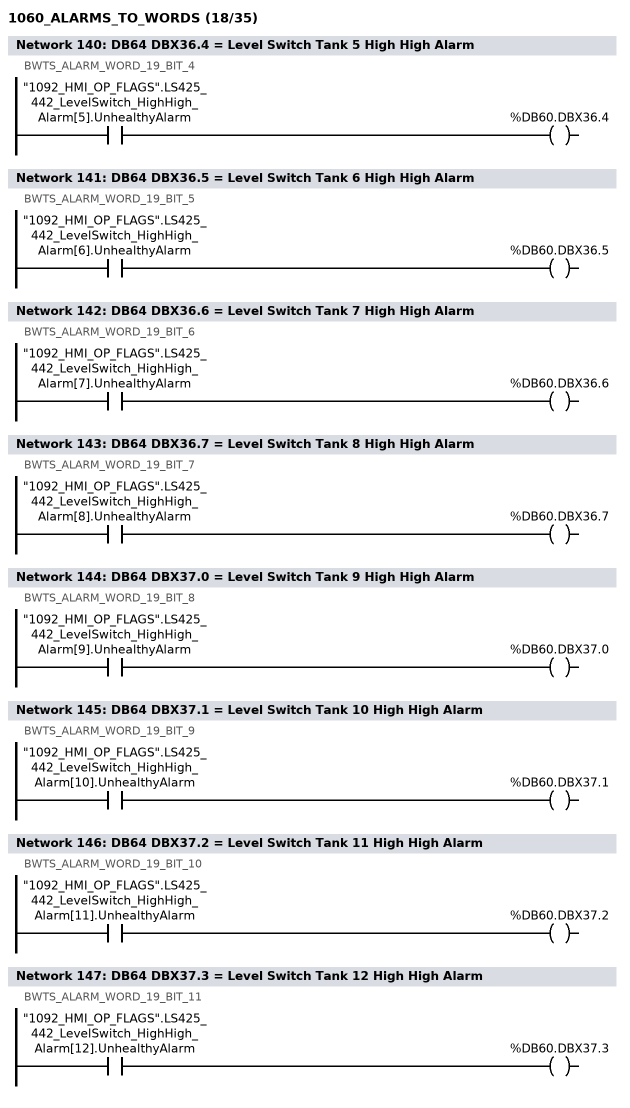
   RUNG wire#powerrail
      Contact( "1092_HMI_OP_FLAGS".LS425_442_LevelSwitch_HighHigh_Alarm[5].UnhealthyAlarm )
      Coil( %DB60.DBX36.4 )
   END_RUNG
   // the same network as SCL:
   %DB60.DBX36.4 := "1092_HMI_OP_FLAGS".LS425_442_LevelSwitch_HighHigh_Alarm[5].UnhealthyAlarm;
END_REGION

REGION Network 141: DB64 DBX36.5 = Level Switch Tank 6 High High Alarm
   // BWTS_ALARM_WORD_19_BIT_5
   RUNG wire#powerrail
      Contact( "1092_HMI_OP_FLAGS".LS425_442_LevelSwitch_HighHigh_Alarm[6].UnhealthyAlarm )
      Coil( %DB60.DBX36.5 )
   END_RUNG
   // the same network as SCL:
   %DB60.DBX36.5 := "1092_HMI_OP_FLAGS".LS425_442_LevelSwitch_HighHigh_Alarm[6].UnhealthyAlarm;
END_REGION

REGION Network 142: DB64 DBX36.6 = Level Switch Tank 7 High High Alarm
   // BWTS_ALARM_WORD_19_BIT_6
   RUNG wire#powerrail
      Contact( "1092_HMI_OP_FLAGS".LS425_442_LevelSwitch_HighHigh_Alarm[7].UnhealthyAlarm )
      Coil( %DB60.DBX36.6 )
   END_RUNG
   // the same network as SCL:
   %DB60.DBX36.6 := "1092_HMI_OP_FLAGS".LS425_442_LevelSwitch_HighHigh_Alarm[7].UnhealthyAlarm;
END_REGION

REGION Network 143: DB64 DBX36.7 = Level Switch Tank 8 High High Alarm
   // BWTS_ALARM_WORD_19_BIT_7
   RUNG wire#powerrail
      Contact( "1092_HMI_OP_FLAGS".LS425_442_LevelSwitch_HighHigh_Alarm[8].UnhealthyAlarm )
      Coil( %DB60.DBX36.7 )
   END_RUNG
   // the same network as SCL:
   %DB60.DBX36.7 := "1092_HMI_OP_FLAGS".LS425_442_LevelSwitch_HighHigh_Alarm[8].UnhealthyAlarm;
END_REGION

REGION Network 144: DB64 DBX37.0 = Level Switch Tank 9 High High Alarm
   // BWTS_ALARM_WORD_19_BIT_8
   RUNG wire#powerrail
      Contact( "1092_HMI_OP_FLAGS".LS425_442_LevelSwitch_HighHigh_Alarm[9].UnhealthyAlarm )
      Coil( %DB60.DBX37.0 )
   END_RUNG
   // the same network as SCL:
   %DB60.DBX37.0 := "1092_HMI_OP_FLAGS".LS425_442_LevelSwitch_HighHigh_Alarm[9].UnhealthyAlarm;
END_REGION

REGION Network 145: DB64 DBX37.1 = Level Switch Tank 10 High High Alarm
   // BWTS_ALARM_WORD_19_BIT_9
   RUNG wire#powerrail
      Contact( "1092_HMI_OP_FLAGS".LS425_442_LevelSwitch_HighHigh_Alarm[10].UnhealthyAlarm )
      Coil( %DB60.DBX37.1 )
   END_RUNG
   // the same network as SCL:
   %DB60.DBX37.1 := "1092_HMI_OP_FLAGS".LS425_442_LevelSwitch_HighHigh_Alarm[10].UnhealthyAlarm;
END_REGION

REGION Network 146: DB64 DBX37.2 = Level Switch Tank 11 High High Alarm
   // BWTS_ALARM_WORD_19_BIT_10
   RUNG wire#powerrail
      Contact( "1092_HMI_OP_FLAGS".LS425_442_LevelSwitch_HighHigh_Alarm[11].UnhealthyAlarm )
      Coil( %DB60.DBX37.2 )
   END_RUNG
   // the same network as SCL:
   %DB60.DBX37.2 := "1092_HMI_OP_FLAGS".LS425_442_LevelSwitch_HighHigh_Alarm[11].UnhealthyAlarm;
END_REGION

REGION Network 147: DB64 DBX37.3 = Level Switch Tank 12 High High Alarm
   // BWTS_ALARM_WORD_19_BIT_11
   RUNG wire#powerrail
      Contact( "1092_HMI_OP_FLAGS".LS425_442_LevelSwitch_HighHigh_Alarm[12].UnhealthyAlarm )
      Coil( %DB60.DBX37.3 )
   END_RUNG
   // the same network as SCL:
   %DB60.DBX37.3 := "1092_HMI_OP_FLAGS".LS425_442_LevelSwitch_HighHigh_Alarm[12].UnhealthyAlarm;
END_REGION

REGION Network 148: DB64 DBX37.4 = Level Switch Tank 13 High High Alarm
   // BWTS_ALARM_WORD_19_BIT_12
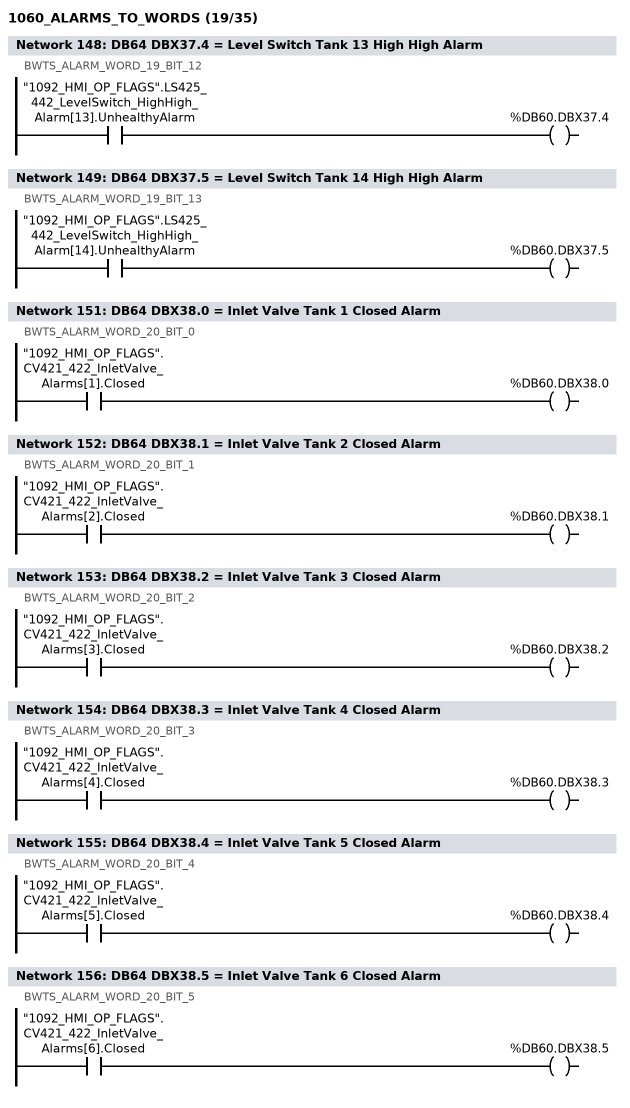
   RUNG wire#powerrail
      Contact( "1092_HMI_OP_FLAGS".LS425_442_LevelSwitch_HighHigh_Alarm[13].UnhealthyAlarm )
      Coil( %DB60.DBX37.4 )
   END_RUNG
   // the same network as SCL:
   %DB60.DBX37.4 := "1092_HMI_OP_FLAGS".LS425_442_LevelSwitch_HighHigh_Alarm[13].UnhealthyAlarm;
END_REGION

REGION Network 149: DB64 DBX37.5 = Level Switch Tank 14 High High Alarm
   // BWTS_ALARM_WORD_19_BIT_13
   RUNG wire#powerrail
      Contact( "1092_HMI_OP_FLAGS".LS425_442_LevelSwitch_HighHigh_Alarm[14].UnhealthyAlarm )
      Coil( %DB60.DBX37.5 )
   END_RUNG
   // the same network as SCL:
   %DB60.DBX37.5 := "1092_HMI_OP_FLAGS".LS425_442_LevelSwitch_HighHigh_Alarm[14].UnhealthyAlarm;
END_REGION

REGION Network 151: DB64 DBX38.0 = Inlet Valve Tank 1 Closed Alarm
   // BWTS_ALARM_WORD_20_BIT_0
   RUNG wire#powerrail
      Contact( "1092_HMI_OP_FLAGS".CV421_422_InletValve_Alarms[1].Closed )
      Coil( %DB60.DBX38.0 )
   END_RUNG
   // the same network as SCL:
   %DB60.DBX38.0 := "1092_HMI_OP_FLAGS".CV421_422_InletValve_Alarms[1].Closed;
END_REGION

REGION Network 152: DB64 DBX38.1 = Inlet Valve Tank 2 Closed Alarm
   // BWTS_ALARM_WORD_20_BIT_1
   RUNG wire#powerrail
      Contact( "1092_HMI_OP_FLAGS".CV421_422_InletValve_Alarms[2].Closed )
      Coil( %DB60.DBX38.1 )
   END_RUNG
   // the same network as SCL:
   %DB60.DBX38.1 := "1092_HMI_OP_FLAGS".CV421_422_InletValve_Alarms[2].Closed;
END_REGION

REGION Network 153: DB64 DBX38.2 = Inlet Valve Tank 3 Closed Alarm
   // BWTS_ALARM_WORD_20_BIT_2
   RUNG wire#powerrail
      Contact( "1092_HMI_OP_FLAGS".CV421_422_InletValve_Alarms[3].Closed )
      Coil( %DB60.DBX38.2 )
   END_RUNG
   // the same network as SCL:
   %DB60.DBX38.2 := "1092_HMI_OP_FLAGS".CV421_422_InletValve_Alarms[3].Closed;
END_REGION

REGION Network 154: DB64 DBX38.3 = Inlet Valve Tank 4 Closed Alarm
   // BWTS_ALARM_WORD_20_BIT_3
   RUNG wire#powerrail
      Contact( "1092_HMI_OP_FLAGS".CV421_422_InletValve_Alarms[4].Closed )
      Coil( %DB60.DBX38.3 )
   END_RUNG
   // the same network as SCL:
   %DB60.DBX38.3 := "1092_HMI_OP_FLAGS".CV421_422_InletValve_Alarms[4].Closed;
END_REGION

REGION Network 155: DB64 DBX38.4 = Inlet Valve Tank 5 Closed Alarm
   // BWTS_ALARM_WORD_20_BIT_4
   RUNG wire#powerrail
      Contact( "1092_HMI_OP_FLAGS".CV421_422_InletValve_Alarms[5].Closed )
      Coil( %DB60.DBX38.4 )
   END_RUNG
   // the same network as SCL:
   %DB60.DBX38.4 := "1092_HMI_OP_FLAGS".CV421_422_InletValve_Alarms[5].Closed;
END_REGION

REGION Network 156: DB64 DBX38.5 = Inlet Valve Tank 6 Closed Alarm
   // BWTS_ALARM_WORD_20_BIT_5
   RUNG wire#powerrail
      Contact( "1092_HMI_OP_FLAGS".CV421_422_InletValve_Alarms[6].Closed )
      Coil( %DB60.DBX38.5 )
   END_RUNG
   // the same network as SCL:
   %DB60.DBX38.5 := "1092_HMI_OP_FLAGS".CV421_422_InletValve_Alarms[6].Closed;
END_REGION

REGION Network 157: DB64 DBX38.6 = Inlet Valve Tank 7 Closed Alarm
   // BWTS_ALARM_WORD_20_BIT_6
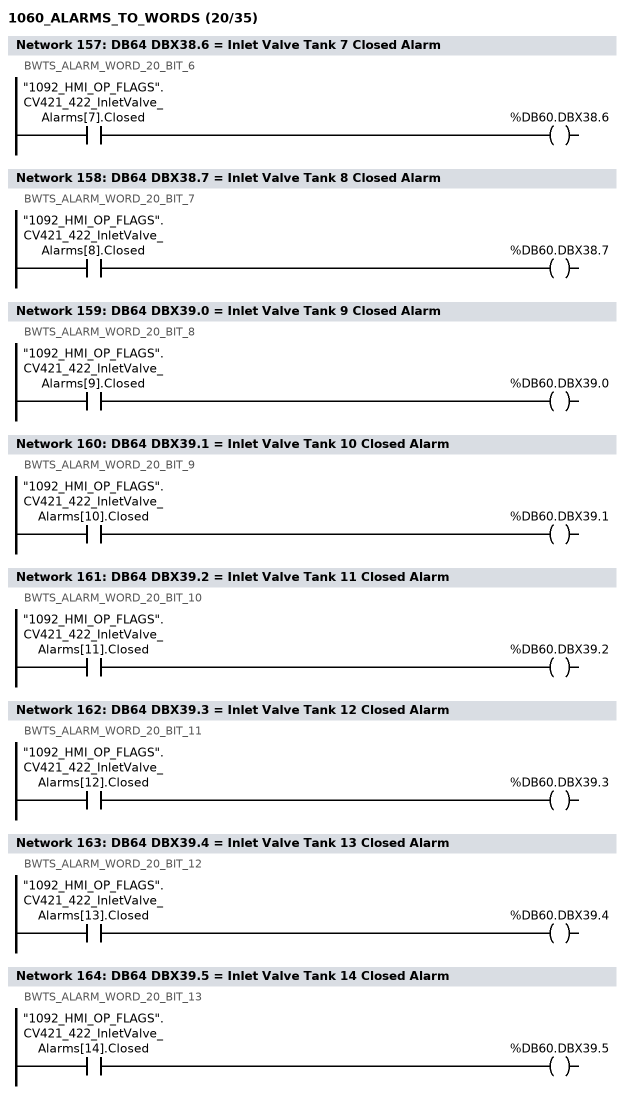
   RUNG wire#powerrail
      Contact( "1092_HMI_OP_FLAGS".CV421_422_InletValve_Alarms[7].Closed )
      Coil( %DB60.DBX38.6 )
   END_RUNG
   // the same network as SCL:
   %DB60.DBX38.6 := "1092_HMI_OP_FLAGS".CV421_422_InletValve_Alarms[7].Closed;
END_REGION

REGION Network 158: DB64 DBX38.7 = Inlet Valve Tank 8 Closed Alarm
   // BWTS_ALARM_WORD_20_BIT_7
   RUNG wire#powerrail
      Contact( "1092_HMI_OP_FLAGS".CV421_422_InletValve_Alarms[8].Closed )
      Coil( %DB60.DBX38.7 )
   END_RUNG
   // the same network as SCL:
   %DB60.DBX38.7 := "1092_HMI_OP_FLAGS".CV421_422_InletValve_Alarms[8].Closed;
END_REGION

REGION Network 159: DB64 DBX39.0 = Inlet Valve Tank 9 Closed Alarm
   // BWTS_ALARM_WORD_20_BIT_8
   RUNG wire#powerrail
      Contact( "1092_HMI_OP_FLAGS".CV421_422_InletValve_Alarms[9].Closed )
      Coil( %DB60.DBX39.0 )
   END_RUNG
   // the same network as SCL:
   %DB60.DBX39.0 := "1092_HMI_OP_FLAGS".CV421_422_InletValve_Alarms[9].Closed;
END_REGION

REGION Network 160: DB64 DBX39.1 = Inlet Valve Tank 10 Closed Alarm
   // BWTS_ALARM_WORD_20_BIT_9
   RUNG wire#powerrail
      Contact( "1092_HMI_OP_FLAGS".CV421_422_InletValve_Alarms[10].Closed )
      Coil( %DB60.DBX39.1 )
   END_RUNG
   // the same network as SCL:
   %DB60.DBX39.1 := "1092_HMI_OP_FLAGS".CV421_422_InletValve_Alarms[10].Closed;
END_REGION

REGION Network 161: DB64 DBX39.2 = Inlet Valve Tank 11 Closed Alarm
   // BWTS_ALARM_WORD_20_BIT_10
   RUNG wire#powerrail
      Contact( "1092_HMI_OP_FLAGS".CV421_422_InletValve_Alarms[11].Closed )
      Coil( %DB60.DBX39.2 )
   END_RUNG
   // the same network as SCL:
   %DB60.DBX39.2 := "1092_HMI_OP_FLAGS".CV421_422_InletValve_Alarms[11].Closed;
END_REGION

REGION Network 162: DB64 DBX39.3 = Inlet Valve Tank 12 Closed Alarm
   // BWTS_ALARM_WORD_20_BIT_11
   RUNG wire#powerrail
      Contact( "1092_HMI_OP_FLAGS".CV421_422_InletValve_Alarms[12].Closed )
      Coil( %DB60.DBX39.3 )
   END_RUNG
   // the same network as SCL:
   %DB60.DBX39.3 := "1092_HMI_OP_FLAGS".CV421_422_InletValve_Alarms[12].Closed;
END_REGION

REGION Network 163: DB64 DBX39.4 = Inlet Valve Tank 13 Closed Alarm
   // BWTS_ALARM_WORD_20_BIT_12
   RUNG wire#powerrail
      Contact( "1092_HMI_OP_FLAGS".CV421_422_InletValve_Alarms[13].Closed )
      Coil( %DB60.DBX39.4 )
   END_RUNG
   // the same network as SCL:
   %DB60.DBX39.4 := "1092_HMI_OP_FLAGS".CV421_422_InletValve_Alarms[13].Closed;
END_REGION

REGION Network 164: DB64 DBX39.5 = Inlet Valve Tank 14 Closed Alarm
   // BWTS_ALARM_WORD_20_BIT_13
   RUNG wire#powerrail
      Contact( "1092_HMI_OP_FLAGS".CV421_422_InletValve_Alarms[14].Closed )
      Coil( %DB60.DBX39.5 )
   END_RUNG
   // the same network as SCL:
   %DB60.DBX39.5 := "1092_HMI_OP_FLAGS".CV421_422_InletValve_Alarms[14].Closed;
END_REGION

REGION Network 166: DB64 DBX40.0 = Inlet Valve Tank 1 Open Alarm
   // BWTS_ALARM_WORD_21_BIT_0
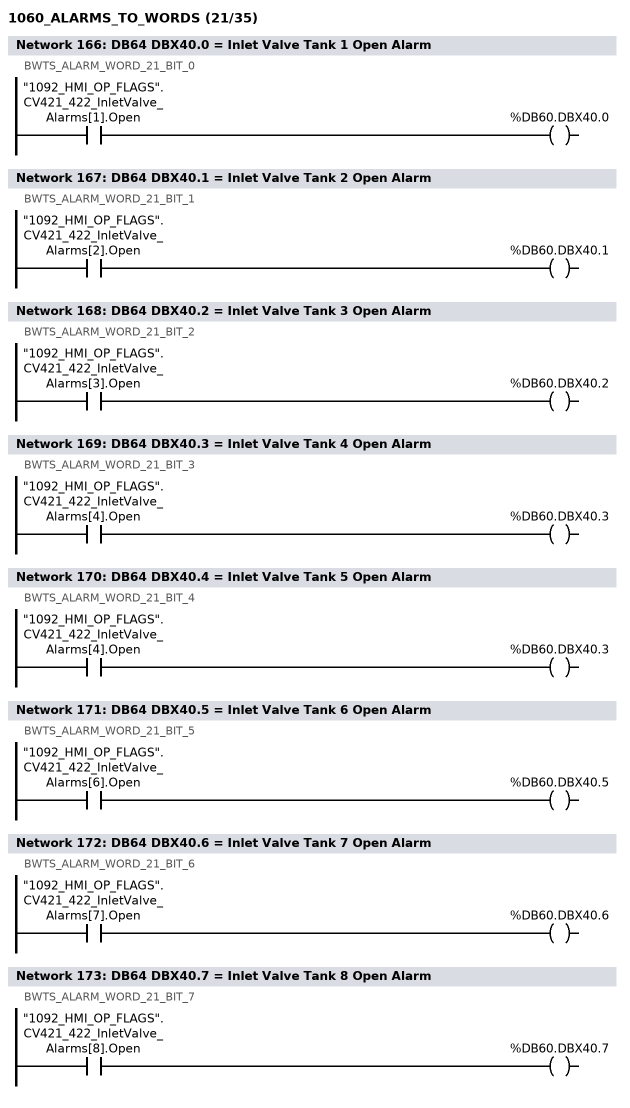
   RUNG wire#powerrail
      Contact( "1092_HMI_OP_FLAGS".CV421_422_InletValve_Alarms[1].Open )
      Coil( %DB60.DBX40.0 )
   END_RUNG
   // the same network as SCL:
   %DB60.DBX40.0 := "1092_HMI_OP_FLAGS".CV421_422_InletValve_Alarms[1].Open;
END_REGION

REGION Network 167: DB64 DBX40.1 = Inlet Valve Tank 2 Open Alarm
   // BWTS_ALARM_WORD_21_BIT_1
   RUNG wire#powerrail
      Contact( "1092_HMI_OP_FLAGS".CV421_422_InletValve_Alarms[2].Open )
      Coil( %DB60.DBX40.1 )
   END_RUNG
   // the same network as SCL:
   %DB60.DBX40.1 := "1092_HMI_OP_FLAGS".CV421_422_InletValve_Alarms[2].Open;
END_REGION

REGION Network 168: DB64 DBX40.2 = Inlet Valve Tank 3 Open Alarm
   // BWTS_ALARM_WORD_21_BIT_2
   RUNG wire#powerrail
      Contact( "1092_HMI_OP_FLAGS".CV421_422_InletValve_Alarms[3].Open )
      Coil( %DB60.DBX40.2 )
   END_RUNG
   // the same network as SCL:
   %DB60.DBX40.2 := "1092_HMI_OP_FLAGS".CV421_422_InletValve_Alarms[3].Open;
END_REGION

REGION Network 169: DB64 DBX40.3 = Inlet Valve Tank 4 Open Alarm
   // BWTS_ALARM_WORD_21_BIT_3
   RUNG wire#powerrail
      Contact( "1092_HMI_OP_FLAGS".CV421_422_InletValve_Alarms[4].Open )
      Coil( %DB60.DBX40.3 )
   END_RUNG
   // the same network as SCL:
   %DB60.DBX40.3 := "1092_HMI_OP_FLAGS".CV421_422_InletValve_Alarms[4].Open;
END_REGION

REGION Network 170: DB64 DBX40.4 = Inlet Valve Tank 5 Open Alarm
   // BWTS_ALARM_WORD_21_BIT_4
   RUNG wire#powerrail
      Contact( "1092_HMI_OP_FLAGS".CV421_422_InletValve_Alarms[4].Open )
      Coil( %DB60.DBX40.3 )
   END_RUNG
   // the same network as SCL:
   %DB60.DBX40.3 := "1092_HMI_OP_FLAGS".CV421_422_InletValve_Alarms[4].Open;
END_REGION

REGION Network 171: DB64 DBX40.5 = Inlet Valve Tank 6 Open Alarm
   // BWTS_ALARM_WORD_21_BIT_5
   RUNG wire#powerrail
      Contact( "1092_HMI_OP_FLAGS".CV421_422_InletValve_Alarms[6].Open )
      Coil( %DB60.DBX40.5 )
   END_RUNG
   // the same network as SCL:
   %DB60.DBX40.5 := "1092_HMI_OP_FLAGS".CV421_422_InletValve_Alarms[6].Open;
END_REGION

REGION Network 172: DB64 DBX40.6 = Inlet Valve Tank 7 Open Alarm
   // BWTS_ALARM_WORD_21_BIT_6
   RUNG wire#powerrail
      Contact( "1092_HMI_OP_FLAGS".CV421_422_InletValve_Alarms[7].Open )
      Coil( %DB60.DBX40.6 )
   END_RUNG
   // the same network as SCL:
   %DB60.DBX40.6 := "1092_HMI_OP_FLAGS".CV421_422_InletValve_Alarms[7].Open;
END_REGION

REGION Network 173: DB64 DBX40.7 = Inlet Valve Tank 8 Open Alarm
   // BWTS_ALARM_WORD_21_BIT_7
   RUNG wire#powerrail
      Contact( "1092_HMI_OP_FLAGS".CV421_422_InletValve_Alarms[8].Open )
      Coil( %DB60.DBX40.7 )
   END_RUNG
   // the same network as SCL:
   %DB60.DBX40.7 := "1092_HMI_OP_FLAGS".CV421_422_InletValve_Alarms[8].Open;
END_REGION

REGION Network 174: DB64 DBX41.0 = Inlet Valve Tank 9 Open Alarm
   // BWTS_ALARM_WORD_21_BIT_8
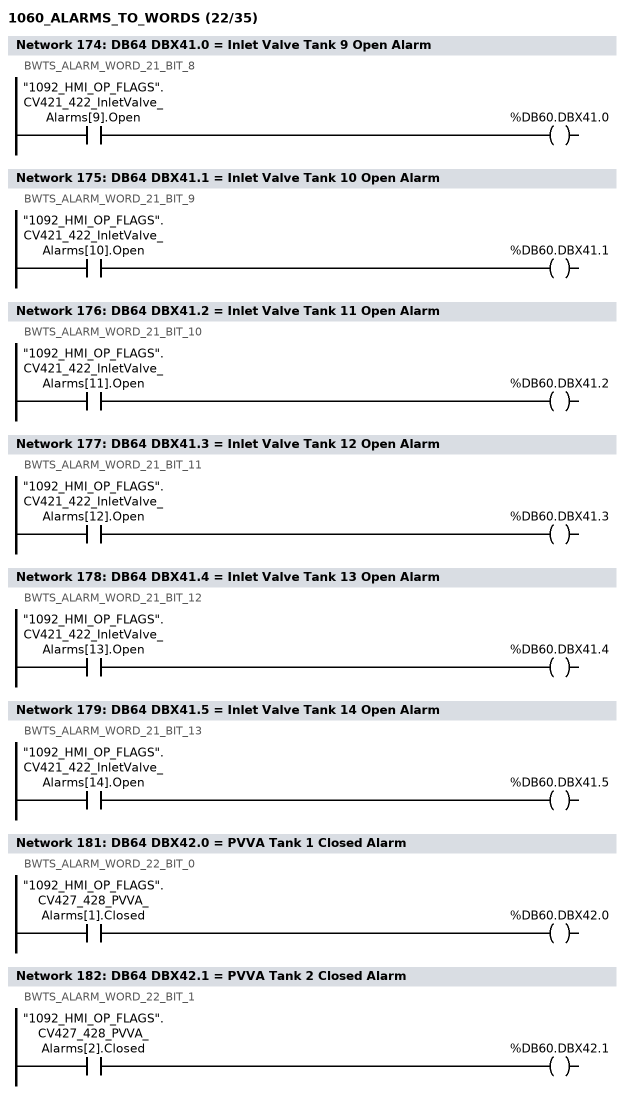
   RUNG wire#powerrail
      Contact( "1092_HMI_OP_FLAGS".CV421_422_InletValve_Alarms[9].Open )
      Coil( %DB60.DBX41.0 )
   END_RUNG
   // the same network as SCL:
   %DB60.DBX41.0 := "1092_HMI_OP_FLAGS".CV421_422_InletValve_Alarms[9].Open;
END_REGION

REGION Network 175: DB64 DBX41.1 = Inlet Valve Tank 10 Open Alarm
   // BWTS_ALARM_WORD_21_BIT_9
   RUNG wire#powerrail
      Contact( "1092_HMI_OP_FLAGS".CV421_422_InletValve_Alarms[10].Open )
      Coil( %DB60.DBX41.1 )
   END_RUNG
   // the same network as SCL:
   %DB60.DBX41.1 := "1092_HMI_OP_FLAGS".CV421_422_InletValve_Alarms[10].Open;
END_REGION

REGION Network 176: DB64 DBX41.2 = Inlet Valve Tank 11 Open Alarm
   // BWTS_ALARM_WORD_21_BIT_10
   RUNG wire#powerrail
      Contact( "1092_HMI_OP_FLAGS".CV421_422_InletValve_Alarms[11].Open )
      Coil( %DB60.DBX41.2 )
   END_RUNG
   // the same network as SCL:
   %DB60.DBX41.2 := "1092_HMI_OP_FLAGS".CV421_422_InletValve_Alarms[11].Open;
END_REGION

REGION Network 177: DB64 DBX41.3 = Inlet Valve Tank 12 Open Alarm
   // BWTS_ALARM_WORD_21_BIT_11
   RUNG wire#powerrail
      Contact( "1092_HMI_OP_FLAGS".CV421_422_InletValve_Alarms[12].Open )
      Coil( %DB60.DBX41.3 )
   END_RUNG
   // the same network as SCL:
   %DB60.DBX41.3 := "1092_HMI_OP_FLAGS".CV421_422_InletValve_Alarms[12].Open;
END_REGION

REGION Network 178: DB64 DBX41.4 = Inlet Valve Tank 13 Open Alarm
   // BWTS_ALARM_WORD_21_BIT_12
   RUNG wire#powerrail
      Contact( "1092_HMI_OP_FLAGS".CV421_422_InletValve_Alarms[13].Open )
      Coil( %DB60.DBX41.4 )
   END_RUNG
   // the same network as SCL:
   %DB60.DBX41.4 := "1092_HMI_OP_FLAGS".CV421_422_InletValve_Alarms[13].Open;
END_REGION

REGION Network 179: DB64 DBX41.5 = Inlet Valve Tank 14 Open Alarm
   // BWTS_ALARM_WORD_21_BIT_13
   RUNG wire#powerrail
      Contact( "1092_HMI_OP_FLAGS".CV421_422_InletValve_Alarms[14].Open )
      Coil( %DB60.DBX41.5 )
   END_RUNG
   // the same network as SCL:
   %DB60.DBX41.5 := "1092_HMI_OP_FLAGS".CV421_422_InletValve_Alarms[14].Open;
END_REGION

REGION Network 181: DB64 DBX42.0 = PVVA Tank 1 Closed Alarm
   // BWTS_ALARM_WORD_22_BIT_0
   RUNG wire#powerrail
      Contact( "1092_HMI_OP_FLAGS".CV427_428_PVVA_Alarms[1].Closed )
      Coil( %DB60.DBX42.0 )
   END_RUNG
   // the same network as SCL:
   %DB60.DBX42.0 := "1092_HMI_OP_FLAGS".CV427_428_PVVA_Alarms[1].Closed;
END_REGION

REGION Network 182: DB64 DBX42.1 = PVVA Tank 2 Closed Alarm
   // BWTS_ALARM_WORD_22_BIT_1
   RUNG wire#powerrail
      Contact( "1092_HMI_OP_FLAGS".CV427_428_PVVA_Alarms[2].Closed )
      Coil( %DB60.DBX42.1 )
   END_RUNG
   // the same network as SCL:
   %DB60.DBX42.1 := "1092_HMI_OP_FLAGS".CV427_428_PVVA_Alarms[2].Closed;
END_REGION

REGION Network 183: DB64 DBX42.2 = PVVA Tank 3 Closed Alarm
   // BWTS_ALARM_WORD_22_BIT_2
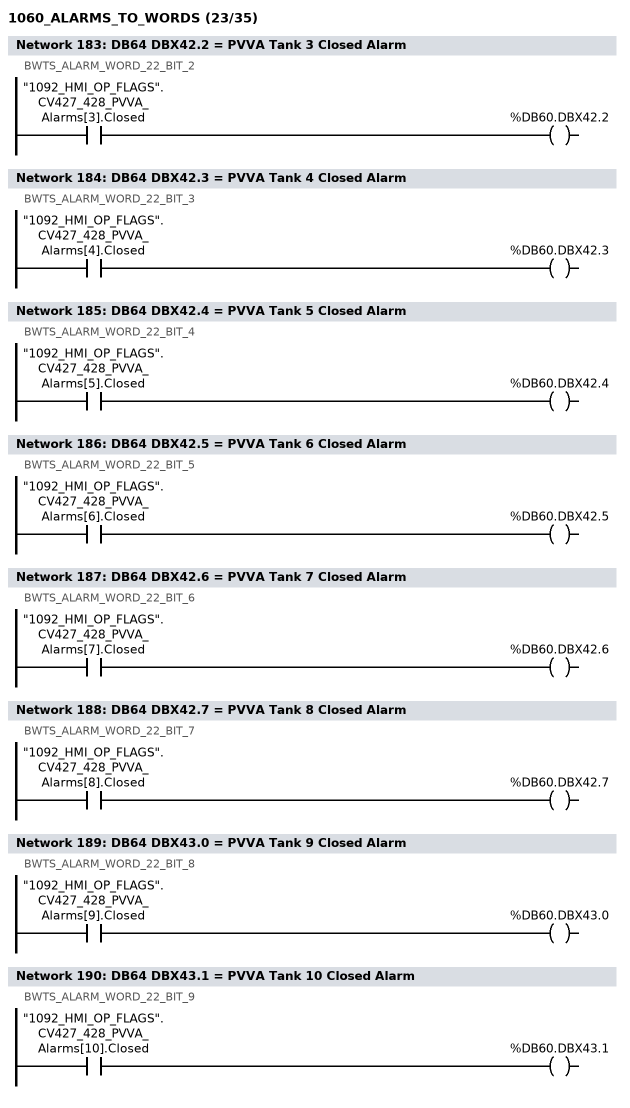
   RUNG wire#powerrail
      Contact( "1092_HMI_OP_FLAGS".CV427_428_PVVA_Alarms[3].Closed )
      Coil( %DB60.DBX42.2 )
   END_RUNG
   // the same network as SCL:
   %DB60.DBX42.2 := "1092_HMI_OP_FLAGS".CV427_428_PVVA_Alarms[3].Closed;
END_REGION

REGION Network 184: DB64 DBX42.3 = PVVA Tank 4 Closed Alarm
   // BWTS_ALARM_WORD_22_BIT_3
   RUNG wire#powerrail
      Contact( "1092_HMI_OP_FLAGS".CV427_428_PVVA_Alarms[4].Closed )
      Coil( %DB60.DBX42.3 )
   END_RUNG
   // the same network as SCL:
   %DB60.DBX42.3 := "1092_HMI_OP_FLAGS".CV427_428_PVVA_Alarms[4].Closed;
END_REGION

REGION Network 185: DB64 DBX42.4 = PVVA Tank 5 Closed Alarm
   // BWTS_ALARM_WORD_22_BIT_4
   RUNG wire#powerrail
      Contact( "1092_HMI_OP_FLAGS".CV427_428_PVVA_Alarms[5].Closed )
      Coil( %DB60.DBX42.4 )
   END_RUNG
   // the same network as SCL:
   %DB60.DBX42.4 := "1092_HMI_OP_FLAGS".CV427_428_PVVA_Alarms[5].Closed;
END_REGION

REGION Network 186: DB64 DBX42.5 = PVVA Tank 6 Closed Alarm
   // BWTS_ALARM_WORD_22_BIT_5
   RUNG wire#powerrail
      Contact( "1092_HMI_OP_FLAGS".CV427_428_PVVA_Alarms[6].Closed )
      Coil( %DB60.DBX42.5 )
   END_RUNG
   // the same network as SCL:
   %DB60.DBX42.5 := "1092_HMI_OP_FLAGS".CV427_428_PVVA_Alarms[6].Closed;
END_REGION

REGION Network 187: DB64 DBX42.6 = PVVA Tank 7 Closed Alarm
   // BWTS_ALARM_WORD_22_BIT_6
   RUNG wire#powerrail
      Contact( "1092_HMI_OP_FLAGS".CV427_428_PVVA_Alarms[7].Closed )
      Coil( %DB60.DBX42.6 )
   END_RUNG
   // the same network as SCL:
   %DB60.DBX42.6 := "1092_HMI_OP_FLAGS".CV427_428_PVVA_Alarms[7].Closed;
END_REGION

REGION Network 188: DB64 DBX42.7 = PVVA Tank 8 Closed Alarm
   // BWTS_ALARM_WORD_22_BIT_7
   RUNG wire#powerrail
      Contact( "1092_HMI_OP_FLAGS".CV427_428_PVVA_Alarms[8].Closed )
      Coil( %DB60.DBX42.7 )
   END_RUNG
   // the same network as SCL:
   %DB60.DBX42.7 := "1092_HMI_OP_FLAGS".CV427_428_PVVA_Alarms[8].Closed;
END_REGION

REGION Network 189: DB64 DBX43.0 = PVVA Tank 9 Closed Alarm
   // BWTS_ALARM_WORD_22_BIT_8
   RUNG wire#powerrail
      Contact( "1092_HMI_OP_FLAGS".CV427_428_PVVA_Alarms[9].Closed )
      Coil( %DB60.DBX43.0 )
   END_RUNG
   // the same network as SCL:
   %DB60.DBX43.0 := "1092_HMI_OP_FLAGS".CV427_428_PVVA_Alarms[9].Closed;
END_REGION

REGION Network 190: DB64 DBX43.1 = PVVA Tank 10 Closed Alarm
   // BWTS_ALARM_WORD_22_BIT_9
   RUNG wire#powerrail
      Contact( "1092_HMI_OP_FLAGS".CV427_428_PVVA_Alarms[10].Closed )
      Coil( %DB60.DBX43.1 )
   END_RUNG
   // the same network as SCL:
   %DB60.DBX43.1 := "1092_HMI_OP_FLAGS".CV427_428_PVVA_Alarms[10].Closed;
END_REGION

REGION Network 191: DB64 DBX43.2 = PVVA Tank 11 Closed Alarm
   // BWTS_ALARM_WORD_22_BIT_10
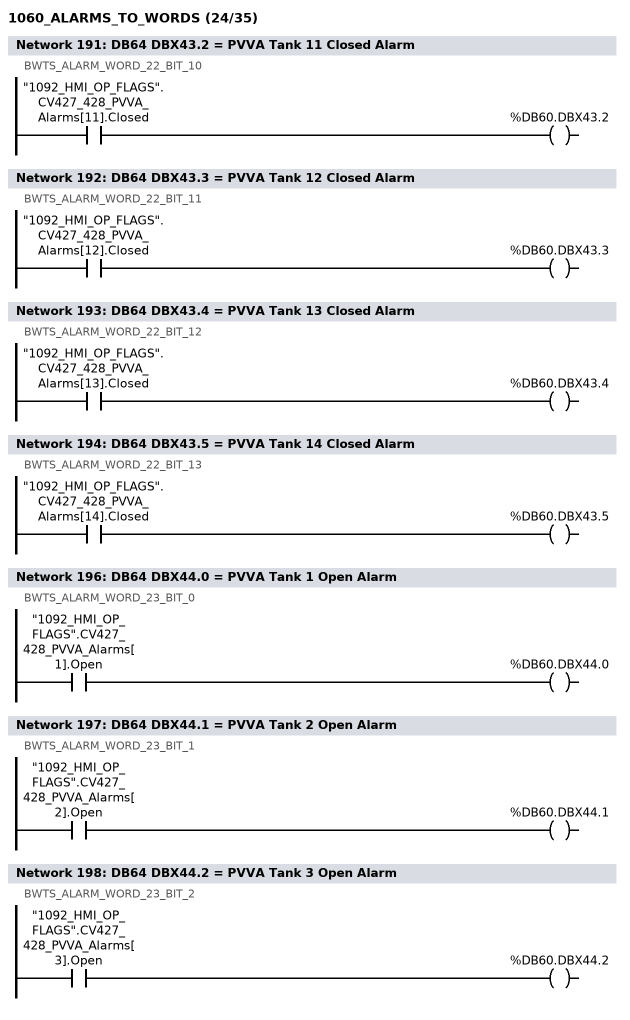
   RUNG wire#powerrail
      Contact( "1092_HMI_OP_FLAGS".CV427_428_PVVA_Alarms[11].Closed )
      Coil( %DB60.DBX43.2 )
   END_RUNG
   // the same network as SCL:
   %DB60.DBX43.2 := "1092_HMI_OP_FLAGS".CV427_428_PVVA_Alarms[11].Closed;
END_REGION

REGION Network 192: DB64 DBX43.3 = PVVA Tank 12 Closed Alarm
   // BWTS_ALARM_WORD_22_BIT_11
   RUNG wire#powerrail
      Contact( "1092_HMI_OP_FLAGS".CV427_428_PVVA_Alarms[12].Closed )
      Coil( %DB60.DBX43.3 )
   END_RUNG
   // the same network as SCL:
   %DB60.DBX43.3 := "1092_HMI_OP_FLAGS".CV427_428_PVVA_Alarms[12].Closed;
END_REGION

REGION Network 193: DB64 DBX43.4 = PVVA Tank 13 Closed Alarm
   // BWTS_ALARM_WORD_22_BIT_12
   RUNG wire#powerrail
      Contact( "1092_HMI_OP_FLAGS".CV427_428_PVVA_Alarms[13].Closed )
      Coil( %DB60.DBX43.4 )
   END_RUNG
   // the same network as SCL:
   %DB60.DBX43.4 := "1092_HMI_OP_FLAGS".CV427_428_PVVA_Alarms[13].Closed;
END_REGION

REGION Network 194: DB64 DBX43.5 = PVVA Tank 14 Closed Alarm
   // BWTS_ALARM_WORD_22_BIT_13
   RUNG wire#powerrail
      Contact( "1092_HMI_OP_FLAGS".CV427_428_PVVA_Alarms[14].Closed )
      Coil( %DB60.DBX43.5 )
   END_RUNG
   // the same network as SCL:
   %DB60.DBX43.5 := "1092_HMI_OP_FLAGS".CV427_428_PVVA_Alarms[14].Closed;
END_REGION

REGION Network 196: DB64 DBX44.0 = PVVA Tank 1 Open Alarm
   // BWTS_ALARM_WORD_23_BIT_0
   RUNG wire#powerrail
      Contact( "1092_HMI_OP_FLAGS".CV427_428_PVVA_Alarms[1].Open )
      Coil( %DB60.DBX44.0 )
   END_RUNG
   // the same network as SCL:
   %DB60.DBX44.0 := "1092_HMI_OP_FLAGS".CV427_428_PVVA_Alarms[1].Open;
END_REGION

REGION Network 197: DB64 DBX44.1 = PVVA Tank 2 Open Alarm
   // BWTS_ALARM_WORD_23_BIT_1
   RUNG wire#powerrail
      Contact( "1092_HMI_OP_FLAGS".CV427_428_PVVA_Alarms[2].Open )
      Coil( %DB60.DBX44.1 )
   END_RUNG
   // the same network as SCL:
   %DB60.DBX44.1 := "1092_HMI_OP_FLAGS".CV427_428_PVVA_Alarms[2].Open;
END_REGION

REGION Network 198: DB64 DBX44.2 = PVVA Tank 3 Open Alarm
   // BWTS_ALARM_WORD_23_BIT_2
   RUNG wire#powerrail
      Contact( "1092_HMI_OP_FLAGS".CV427_428_PVVA_Alarms[3].Open )
      Coil( %DB60.DBX44.2 )
   END_RUNG
   // the same network as SCL:
   %DB60.DBX44.2 := "1092_HMI_OP_FLAGS".CV427_428_PVVA_Alarms[3].Open;
END_REGION

REGION Network 199: DB64 DBX44.3 = PVVA Tank 4 Open Alarm
   // BWTS_ALARM_WORD_23_BIT_3
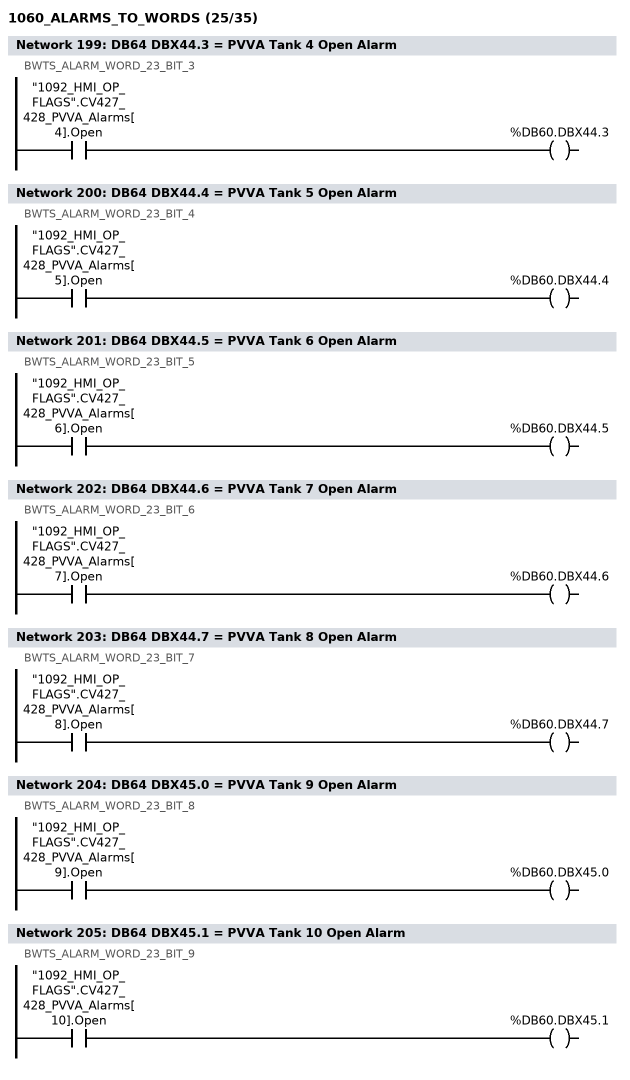
   RUNG wire#powerrail
      Contact( "1092_HMI_OP_FLAGS".CV427_428_PVVA_Alarms[4].Open )
      Coil( %DB60.DBX44.3 )
   END_RUNG
   // the same network as SCL:
   %DB60.DBX44.3 := "1092_HMI_OP_FLAGS".CV427_428_PVVA_Alarms[4].Open;
END_REGION

REGION Network 200: DB64 DBX44.4 = PVVA Tank 5 Open Alarm
   // BWTS_ALARM_WORD_23_BIT_4
   RUNG wire#powerrail
      Contact( "1092_HMI_OP_FLAGS".CV427_428_PVVA_Alarms[5].Open )
      Coil( %DB60.DBX44.4 )
   END_RUNG
   // the same network as SCL:
   %DB60.DBX44.4 := "1092_HMI_OP_FLAGS".CV427_428_PVVA_Alarms[5].Open;
END_REGION

REGION Network 201: DB64 DBX44.5 = PVVA Tank 6 Open Alarm
   // BWTS_ALARM_WORD_23_BIT_5
   RUNG wire#powerrail
      Contact( "1092_HMI_OP_FLAGS".CV427_428_PVVA_Alarms[6].Open )
      Coil( %DB60.DBX44.5 )
   END_RUNG
   // the same network as SCL:
   %DB60.DBX44.5 := "1092_HMI_OP_FLAGS".CV427_428_PVVA_Alarms[6].Open;
END_REGION

REGION Network 202: DB64 DBX44.6 = PVVA Tank 7 Open Alarm
   // BWTS_ALARM_WORD_23_BIT_6
   RUNG wire#powerrail
      Contact( "1092_HMI_OP_FLAGS".CV427_428_PVVA_Alarms[7].Open )
      Coil( %DB60.DBX44.6 )
   END_RUNG
   // the same network as SCL:
   %DB60.DBX44.6 := "1092_HMI_OP_FLAGS".CV427_428_PVVA_Alarms[7].Open;
END_REGION
